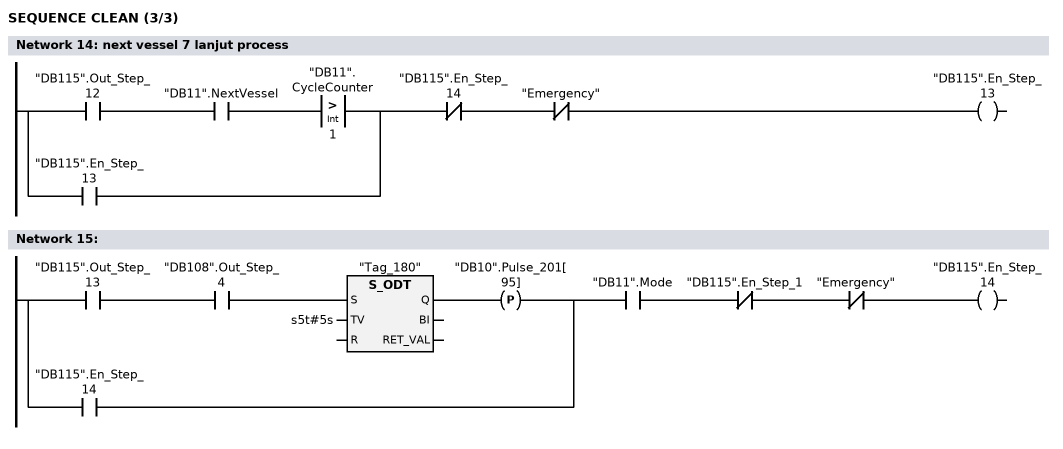
   RUNG wire#powerrail
      Contact( "DB115".Out_Step_12 )
      Contact( "DB11".NextVessel )
      { S7_Templates := "SrcType := Int" } GT_Contact(in1 := "DB11".CycleCounter, in2 := 1)
      wire#w1
      I_Contact( "DB115".En_Step_14 )
      I_Contact( "Emergency" )
      Coil( "DB115".En_Step_13 )
   END_RUNG
   RUNG wire#powerrail
      Contact( "DB115".En_Step_13 )
   END_RUNG wire#w1
   // the same network as SCL:
   "DB115".En_Step_13 := (("DB115".Out_Step_12 AND "DB11".NextVessel AND ("DB11".CycleCounter > 1)) OR "DB115".En_Step_13) AND NOT "DB115".En_Step_14 AND NOT "Emergency";
END_REGION

REGION Network 15
   RUNG wire#powerrail
      Contact( "DB115".Out_Step_13 )
      Contact( "DB108".Out_Step_4 )
      S_ODT(T_NO := "Tag_180", TV := s5t#5s, R :=, BI =>, RET_VAL =>)
      P_Trig( "DB10".Pulse_201[95] )
      wire#w1
      Contact( "DB11".Mode )
      I_Contact( "DB115".En_Step_1 )
      I_Contact( "Emergency" )
      Coil( "DB115".En_Step_14 )
   END_RUNG
   RUNG wire#powerrail
      Contact( "DB115".En_Step_14 )
   END_RUNG wire#w1
   // the same network as SCL:
   #_s5time1 := S_ODT(T_NO := "Tag_180",
                      S := "DB115".Out_Step_13 AND "DB108".Out_Step_4,
                      TV := s5t#5s,
                      Q => #_w1);
   #_w2 := #_w1 AND NOT "DB10".Pulse_201[95];   // rising edge
   "DB10".Pulse_201[95] := #_w1;
   "DB115".En_Step_14 := (#_w2 OR "DB115".En_Step_14) AND "DB11".Mode AND NOT "DB115".En_Step_1 AND NOT "Emergency";
END_REGION
END_FUNCTION

FUNCTION "SEQUENCE CYCLE" : Void   // FC36, LAD
{ S7_Optimized_Access := 'TRUE' }
VERSION : 0.1
   VAR_TEMP   // added for the SCL form of the ladder/FBD networks
      _w1 : Bool;
      _w2 : Bool;
      _w3 : Bool;
      _s5time1 : S5Time;
      _w4 : Bool;
      _w5 : Bool;
   END_VAR
BEGIN

REGION Network 1: Dari supply ke vessel 1
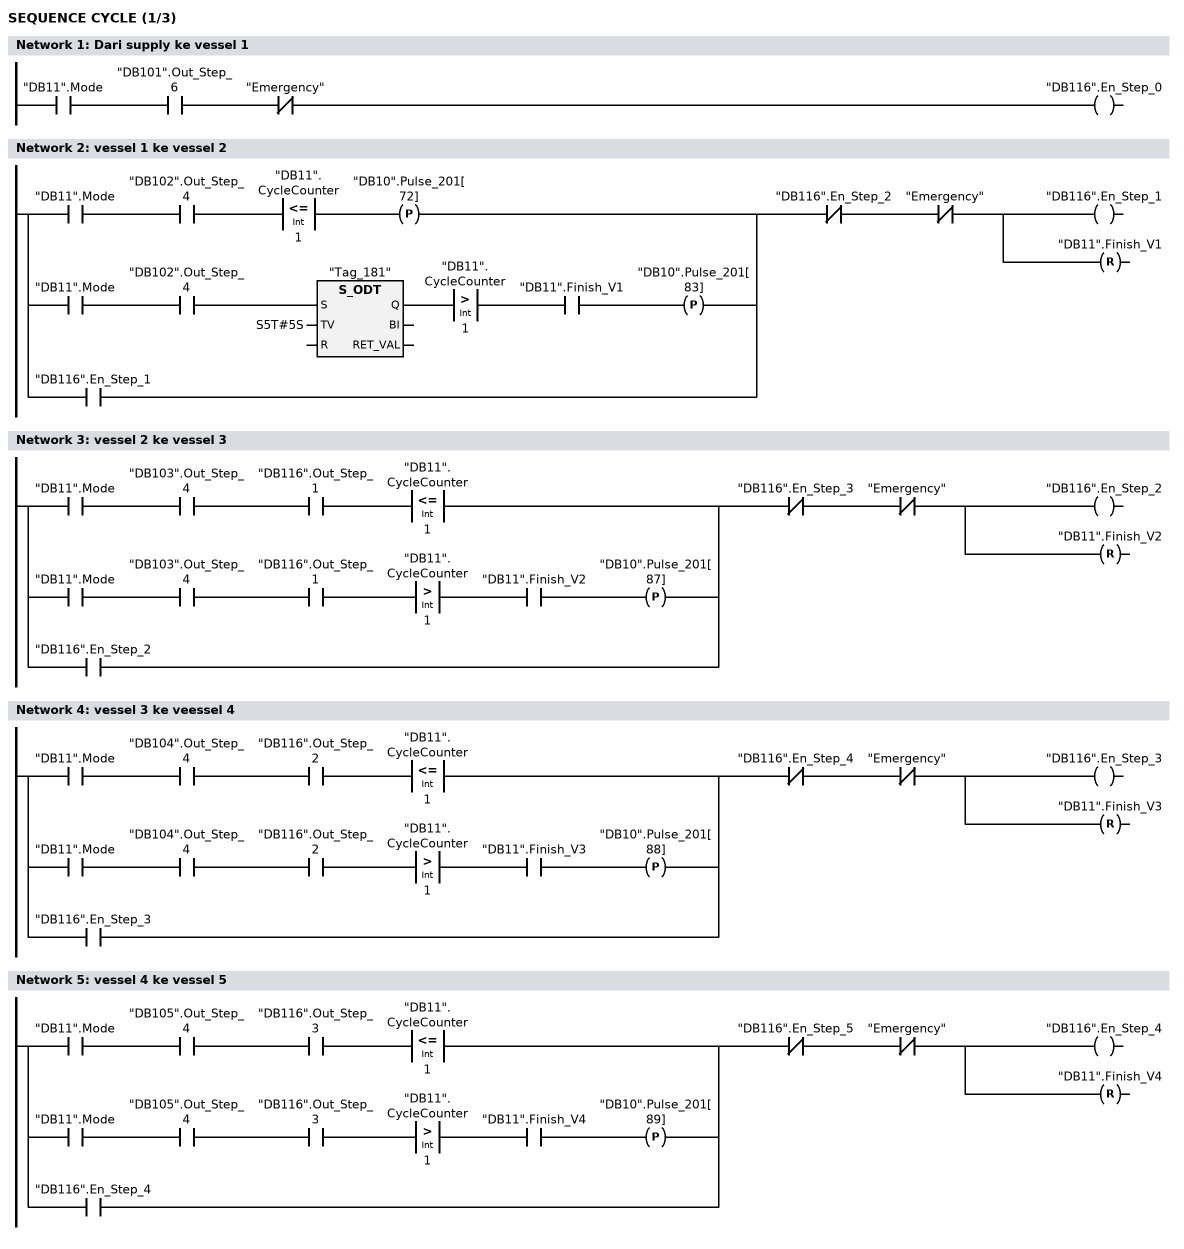
   RUNG wire#powerrail
      Contact( "DB11".Mode )
      Contact( "DB101".Out_Step_6 )
      I_Contact( "Emergency" )
      Coil( "DB116".En_Step_0 )
   END_RUNG
   // the same network as SCL:
   "DB116".En_Step_0 := "DB11".Mode AND "DB101".Out_Step_6 AND NOT "Emergency";
END_REGION

REGION Network 2: vessel 1 ke vessel 2
   RUNG wire#powerrail
      Contact( "DB11".Mode )
      Contact( "DB102".Out_Step_4 )
      { S7_Templates := "SrcType := Int" } LE_Contact(in1 := "DB11".CycleCounter, in2 := 1)
      P_Trig( "DB10".Pulse_201[72] )
      wire#w1
      I_Contact( "DB116".En_Step_2 )
      I_Contact( "Emergency" )
      wire#w2
      Coil( "DB116".En_Step_1 )
   END_RUNG
   RUNG wire#powerrail
      Contact( "DB11".Mode )
      Contact( "DB102".Out_Step_4 )
      S_ODT(T_NO := "Tag_181", TV := S5T#5S, R :=, BI =>, RET_VAL =>)
      { S7_Templates := "SrcType := Int" } GT_Contact(in1 := "DB11".CycleCounter, in2 := 1)
      Contact( "DB11".Finish_V1 )
      P_Trig( "DB10".Pulse_201[83] )
   END_RUNG wire#w1
   RUNG wire#powerrail
      Contact( "DB116".En_Step_1 )
   END_RUNG wire#w1
   RUNG wire#w2
      R_Coil( "DB11".Finish_V1 )
   END_RUNG
   // the same network as SCL:
   #_w1 := "DB11".Mode AND "DB102".Out_Step_4 AND ("DB11".CycleCounter <= 1);
   #_w2 := #_w1 AND NOT "DB10".Pulse_201[72];   // rising edge
   "DB10".Pulse_201[72] := #_w1;
   #_s5time1 := S_ODT(T_NO := "Tag_181", S := "DB11".Mode AND "DB102".Out_Step_4, TV := S5T#5S, Q => #_w3);
   #_w4 := #_w3 AND ("DB11".CycleCounter > 1) AND "DB11".Finish_V1;
   #_w5 := #_w4 AND NOT "DB10".Pulse_201[83];   // rising edge
   "DB10".Pulse_201[83] := #_w4;
   "DB116".En_Step_1 := (#_w2 OR #_w5 OR "DB116".En_Step_1) AND NOT "DB116".En_Step_2 AND NOT "Emergency";
   IF "DB116".En_Step_1 THEN "DB11".Finish_V1 := FALSE; END_IF;
END_REGION

REGION Network 3: vessel 2 ke vessel 3
   RUNG wire#powerrail
      Contact( "DB11".Mode )
      Contact( "DB103".Out_Step_4 )
      Contact( "DB116".Out_Step_1 )
      { S7_Templates := "SrcType := Int" } LE_Contact(in1 := "DB11".CycleCounter, in2 := 1)
      wire#w1
      I_Contact( "DB116".En_Step_3 )
      I_Contact( "Emergency" )
      wire#w2
      Coil( "DB116".En_Step_2 )
   END_RUNG
   RUNG wire#powerrail
      Contact( "DB11".Mode )
      Contact( "DB103".Out_Step_4 )
      Contact( "DB116".Out_Step_1 )
      { S7_Templates := "SrcType := Int" } GT_Contact(in1 := "DB11".CycleCounter, in2 := 1)
      Contact( "DB11".Finish_V2 )
      P_Trig( "DB10".Pulse_201[87] )
   END_RUNG wire#w1
   RUNG wire#powerrail
      Contact( "DB116".En_Step_2 )
   END_RUNG wire#w1
   RUNG wire#w2
      R_Coil( "DB11".Finish_V2 )
   END_RUNG
   // the same network as SCL:
   #_w1 := "DB11".Mode AND "DB103".Out_Step_4 AND "DB116".Out_Step_1 AND ("DB11".CycleCounter > 1) AND "DB11".Finish_V2;
   #_w2 := #_w1 AND NOT "DB10".Pulse_201[87];   // rising edge
   "DB10".Pulse_201[87] := #_w1;
   "DB116".En_Step_2 := (("DB11".Mode AND "DB103".Out_Step_4 AND "DB116".Out_Step_1 AND ("DB11".CycleCounter <= 1)) OR #_w2 OR "DB116".En_Step_2) AND NOT "DB116".En_Step_3 AND NOT "Emergency";
   IF "DB116".En_Step_2 THEN "DB11".Finish_V2 := FALSE; END_IF;
END_REGION

REGION Network 4: vessel 3 ke veessel 4
   RUNG wire#powerrail
      Contact( "DB11".Mode )
      Contact( "DB104".Out_Step_4 )
      Contact( "DB116".Out_Step_2 )
      { S7_Templates := "SrcType := Int" } LE_Contact(in1 := "DB11".CycleCounter, in2 := 1)
      wire#w1
      I_Contact( "DB116".En_Step_4 )
      I_Contact( "Emergency" )
      wire#w2
      Coil( "DB116".En_Step_3 )
   END_RUNG
   RUNG wire#powerrail
      Contact( "DB11".Mode )
      Contact( "DB104".Out_Step_4 )
      Contact( "DB116".Out_Step_2 )
      { S7_Templates := "SrcType := Int" } GT_Contact(in1 := "DB11".CycleCounter, in2 := 1)
      Contact( "DB11".Finish_V3 )
      P_Trig( "DB10".Pulse_201[88] )
   END_RUNG wire#w1
   RUNG wire#powerrail
      Contact( "DB116".En_Step_3 )
   END_RUNG wire#w1
   RUNG wire#w2
      R_Coil( "DB11".Finish_V3 )
   END_RUNG
   // the same network as SCL:
   #_w1 := "DB11".Mode AND "DB104".Out_Step_4 AND "DB116".Out_Step_2 AND ("DB11".CycleCounter > 1) AND "DB11".Finish_V3;
   #_w2 := #_w1 AND NOT "DB10".Pulse_201[88];   // rising edge
   "DB10".Pulse_201[88] := #_w1;
   "DB116".En_Step_3 := (("DB11".Mode AND "DB104".Out_Step_4 AND "DB116".Out_Step_2 AND ("DB11".CycleCounter <= 1)) OR #_w2 OR "DB116".En_Step_3) AND NOT "DB116".En_Step_4 AND NOT "Emergency";
   IF "DB116".En_Step_3 THEN "DB11".Finish_V3 := FALSE; END_IF;
END_REGION

REGION Network 5: vessel 4 ke vessel 5
   RUNG wire#powerrail
      Contact( "DB11".Mode )
      Contact( "DB105".Out_Step_4 )
      Contact( "DB116".Out_Step_3 )
      { S7_Templates := "SrcType := Int" } LE_Contact(in1 := "DB11".CycleCounter, in2 := 1)
      wire#w1
      I_Contact( "DB116".En_Step_5 )
      I_Contact( "Emergency" )
      wire#w2
      Coil( "DB116".En_Step_4 )
   END_RUNG
   RUNG wire#powerrail
      Contact( "DB11".Mode )
      Contact( "DB105".Out_Step_4 )
      Contact( "DB116".Out_Step_3 )
      { S7_Templates := "SrcType := Int" } GT_Contact(in1 := "DB11".CycleCounter, in2 := 1)
      Contact( "DB11".Finish_V4 )
      P_Trig( "DB10".Pulse_201[89] )
   END_RUNG wire#w1
   RUNG wire#powerrail
      Contact( "DB116".En_Step_4 )
   END_RUNG wire#w1
   RUNG wire#w2
      R_Coil( "DB11".Finish_V4 )
   END_RUNG
   // the same network as SCL:
   #_w1 := "DB11".Mode AND "DB105".Out_Step_4 AND "DB116".Out_Step_3 AND ("DB11".CycleCounter > 1) AND "DB11".Finish_V4;
   #_w2 := #_w1 AND NOT "DB10".Pulse_201[89];   // rising edge
   "DB10".Pulse_201[89] := #_w1;
   "DB116".En_Step_4 := (("DB11".Mode AND "DB105".Out_Step_4 AND "DB116".Out_Step_3 AND ("DB11".CycleCounter <= 1)) OR #_w2 OR "DB116".En_Step_4) AND NOT "DB116".En_Step_5 AND NOT "Emergency";
   IF "DB116".En_Step_4 THEN "DB11".Finish_V4 := FALSE; END_IF;
END_REGION

REGION Network 6: vessel 5 ke vessel 6
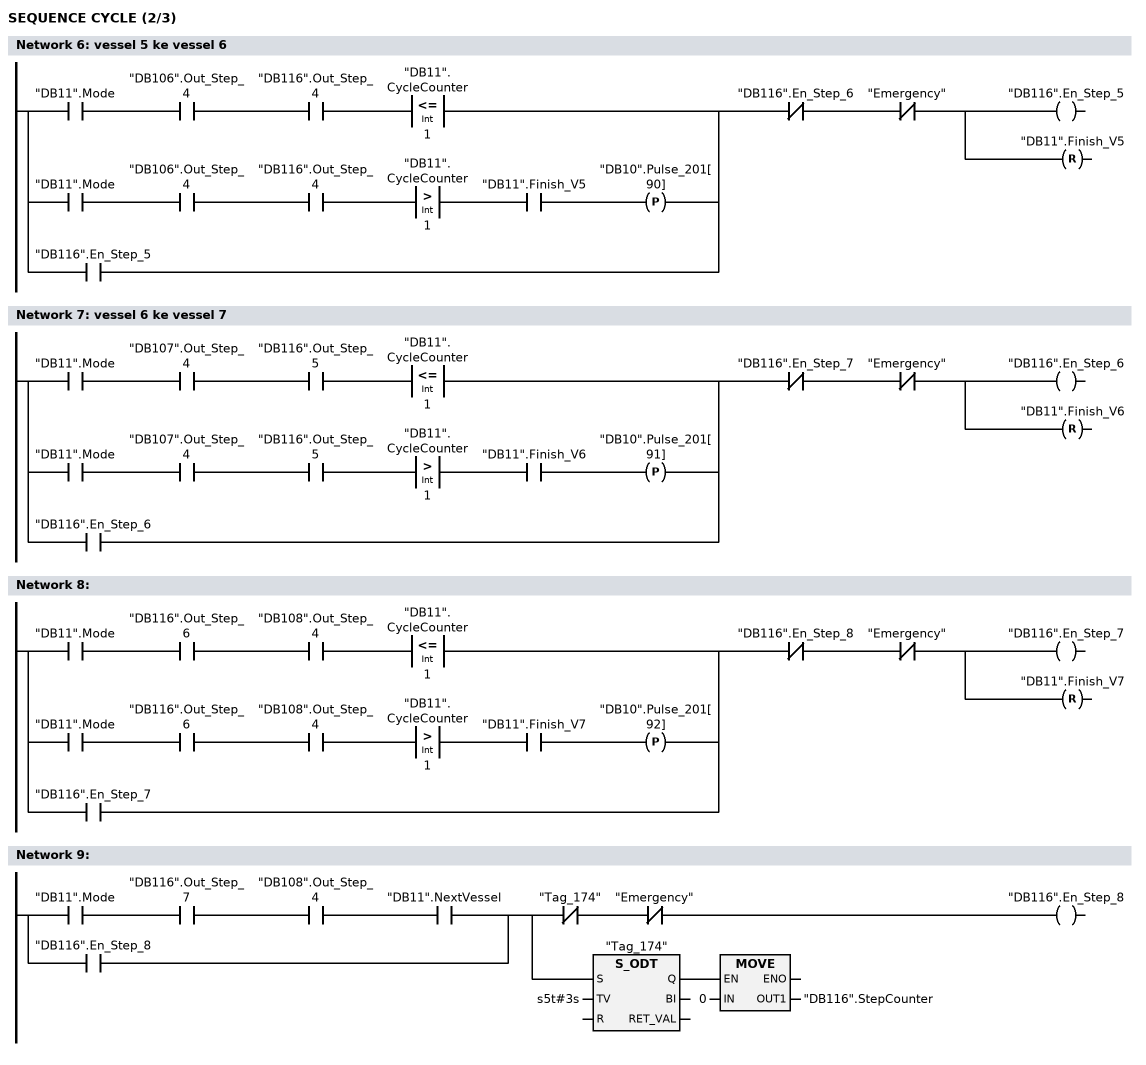
   RUNG wire#powerrail
      Contact( "DB11".Mode )
      Contact( "DB106".Out_Step_4 )
      Contact( "DB116".Out_Step_4 )
      { S7_Templates := "SrcType := Int" } LE_Contact(in1 := "DB11".CycleCounter, in2 := 1)
      wire#w1
      I_Contact( "DB116".En_Step_6 )
      I_Contact( "Emergency" )
      wire#w2
      Coil( "DB116".En_Step_5 )
   END_RUNG
   RUNG wire#powerrail
      Contact( "DB11".Mode )
      Contact( "DB106".Out_Step_4 )
      Contact( "DB116".Out_Step_4 )
      { S7_Templates := "SrcType := Int" } GT_Contact(in1 := "DB11".CycleCounter, in2 := 1)
      Contact( "DB11".Finish_V5 )
      P_Trig( "DB10".Pulse_201[90] )
   END_RUNG wire#w1
   RUNG wire#powerrail
      Contact( "DB116".En_Step_5 )
   END_RUNG wire#w1
   RUNG wire#w2
      R_Coil( "DB11".Finish_V5 )
   END_RUNG
   // the same network as SCL:
   #_w1 := "DB11".Mode AND "DB106".Out_Step_4 AND "DB116".Out_Step_4 AND ("DB11".CycleCounter > 1) AND "DB11".Finish_V5;
   #_w2 := #_w1 AND NOT "DB10".Pulse_201[90];   // rising edge
   "DB10".Pulse_201[90] := #_w1;
   "DB116".En_Step_5 := (("DB11".Mode AND "DB106".Out_Step_4 AND "DB116".Out_Step_4 AND ("DB11".CycleCounter <= 1)) OR #_w2 OR "DB116".En_Step_5) AND NOT "DB116".En_Step_6 AND NOT "Emergency";
   IF "DB116".En_Step_5 THEN "DB11".Finish_V5 := FALSE; END_IF;
END_REGION

REGION Network 7: vessel 6 ke vessel 7
   RUNG wire#powerrail
      Contact( "DB11".Mode )
      Contact( "DB107".Out_Step_4 )
      Contact( "DB116".Out_Step_5 )
      { S7_Templates := "SrcType := Int" } LE_Contact(in1 := "DB11".CycleCounter, in2 := 1)
      wire#w1
      I_Contact( "DB116".En_Step_7 )
      I_Contact( "Emergency" )
      wire#w2
      Coil( "DB116".En_Step_6 )
   END_RUNG
   RUNG wire#powerrail
      Contact( "DB11".Mode )
      Contact( "DB107".Out_Step_4 )
      Contact( "DB116".Out_Step_5 )
      { S7_Templates := "SrcType := Int" } GT_Contact(in1 := "DB11".CycleCounter, in2 := 1)
      Contact( "DB11".Finish_V6 )
      P_Trig( "DB10".Pulse_201[91] )
   END_RUNG wire#w1
   RUNG wire#powerrail
      Contact( "DB116".En_Step_6 )
   END_RUNG wire#w1
   RUNG wire#w2
      R_Coil( "DB11".Finish_V6 )
   END_RUNG
   // the same network as SCL:
   #_w1 := "DB11".Mode AND "DB107".Out_Step_4 AND "DB116".Out_Step_5 AND ("DB11".CycleCounter > 1) AND "DB11".Finish_V6;
   #_w2 := #_w1 AND NOT "DB10".Pulse_201[91];   // rising edge
   "DB10".Pulse_201[91] := #_w1;
   "DB116".En_Step_6 := (("DB11".Mode AND "DB107".Out_Step_4 AND "DB116".Out_Step_5 AND ("DB11".CycleCounter <= 1)) OR #_w2 OR "DB116".En_Step_6) AND NOT "DB116".En_Step_7 AND NOT "Emergency";
   IF "DB116".En_Step_6 THEN "DB11".Finish_V6 := FALSE; END_IF;
END_REGION

REGION Network 8
   RUNG wire#powerrail
      Contact( "DB11".Mode )
      Contact( "DB116".Out_Step_6 )
      Contact( "DB108".Out_Step_4 )
      { S7_Templates := "SrcType := Int" } LE_Contact(in1 := "DB11".CycleCounter, in2 := 1)
      wire#w1
      I_Contact( "DB116".En_Step_8 )
      I_Contact( "Emergency" )
      wire#w2
      Coil( "DB116".En_Step_7 )
   END_RUNG
   RUNG wire#powerrail
      Contact( "DB11".Mode )
      Contact( "DB116".Out_Step_6 )
      Contact( "DB108".Out_Step_4 )
      { S7_Templates := "SrcType := Int" } GT_Contact(in1 := "DB11".CycleCounter, in2 := 1)
      Contact( "DB11".Finish_V7 )
      P_Trig( "DB10".Pulse_201[92] )
   END_RUNG wire#w1
   RUNG wire#powerrail
      Contact( "DB116".En_Step_7 )
   END_RUNG wire#w1
   RUNG wire#w2
      R_Coil( "DB11".Finish_V7 )
   END_RUNG
   // the same network as SCL:
   #_w1 := "DB11".Mode AND "DB116".Out_Step_6 AND "DB108".Out_Step_4 AND ("DB11".CycleCounter > 1) AND "DB11".Finish_V7;
   #_w2 := #_w1 AND NOT "DB10".Pulse_201[92];   // rising edge
   "DB10".Pulse_201[92] := #_w1;
   "DB116".En_Step_7 := (("DB11".Mode AND "DB116".Out_Step_6 AND "DB108".Out_Step_4 AND ("DB11".CycleCounter <= 1)) OR #_w2 OR "DB116".En_Step_7) AND NOT "DB116".En_Step_8 AND NOT "Emergency";
   IF "DB116".En_Step_7 THEN "DB11".Finish_V7 := FALSE; END_IF;
END_REGION

REGION Network 9
   RUNG wire#powerrail
      Contact( "DB11".Mode )
      Contact( "DB116".Out_Step_7 )
      Contact( "DB108".Out_Step_4 )
      Contact( "DB11".NextVessel )
      wire#w1
      I_Contact( "Tag_174" )
      I_Contact( "Emergency" )
      Coil( "DB116".En_Step_8 )
   END_RUNG
   RUNG wire#powerrail
      Contact( "DB116".En_Step_8 )
   END_RUNG wire#w1
   RUNG wire#w1
      S_ODT(T_NO := "Tag_174", TV := s5t#3s, R :=, BI =>, RET_VAL =>)
      Move(in := 0, out1 => "DB116".StepCounter)
   END_RUNG
   // the same network as SCL:
   #_w1 := ("DB11".Mode AND "DB116".Out_Step_7 AND "DB108".Out_Step_4 AND "DB11".NextVessel) OR "DB116".En_Step_8;
   "DB116".En_Step_8 := #_w1 AND NOT "Tag_174" AND NOT "Emergency";
   #_s5time1 := S_ODT(T_NO := "Tag_174", S := #_w1, TV := s5t#3s, Q => #_w2);
   IF #_w2 THEN "DB116".StepCounter := 0; END_IF;
END_REGION

REGION Network 10
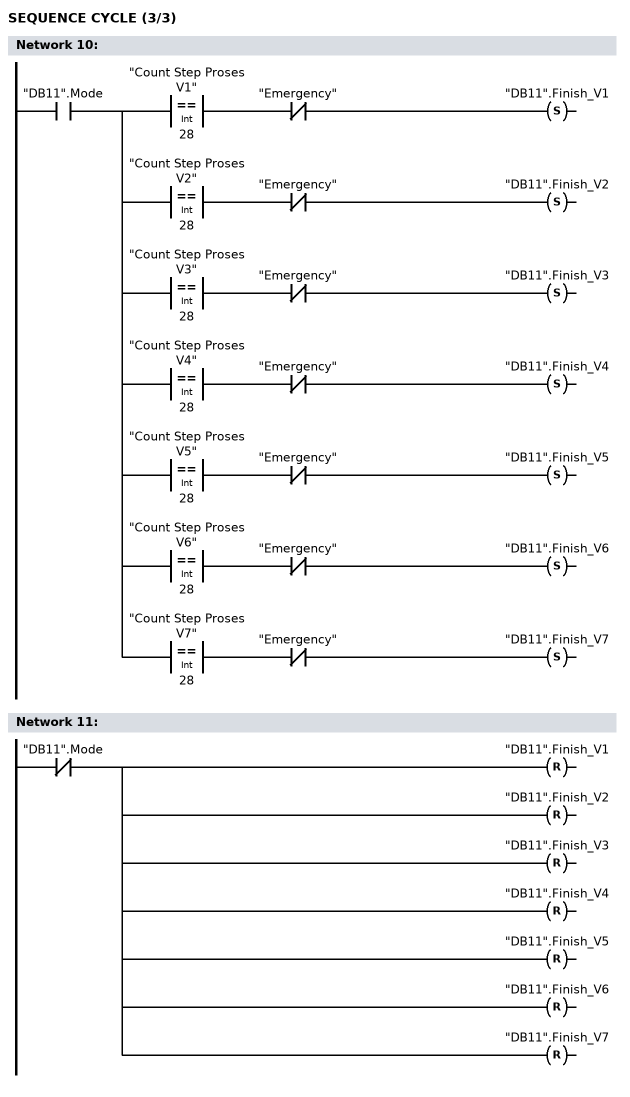
   RUNG wire#powerrail
      Contact( "DB11".Mode )
      wire#w1
      { S7_Templates := "SrcType := Int" } EQ_Contact(in1 := "Count Step Proses V1", in2 := 28)
      I_Contact( "Emergency" )
      S_Coil( "DB11".Finish_V1 )
   END_RUNG
   RUNG wire#w1
      { S7_Templates := "SrcType := Int" } EQ_Contact(in1 := "Count Step Proses V2", in2 := 28)
      I_Contact( "Emergency" )
      S_Coil( "DB11".Finish_V2 )
   END_RUNG
   RUNG wire#w1
      { S7_Templates := "SrcType := Int" } EQ_Contact(in1 := "Count Step Proses V3", in2 := 28)
      I_Contact( "Emergency" )
      S_Coil( "DB11".Finish_V3 )
   END_RUNG
   RUNG wire#w1
      { S7_Templates := "SrcType := Int" } EQ_Contact(in1 := "Count Step Proses V4", in2 := 28)
      I_Contact( "Emergency" )
      S_Coil( "DB11".Finish_V4 )
   END_RUNG
   RUNG wire#w1
      { S7_Templates := "SrcType := Int" } EQ_Contact(in1 := "Count Step Proses V5", in2 := 28)
      I_Contact( "Emergency" )
      S_Coil( "DB11".Finish_V5 )
   END_RUNG
   RUNG wire#w1
      { S7_Templates := "SrcType := Int" } EQ_Contact(in1 := "Count Step Proses V6", in2 := 28)
      I_Contact( "Emergency" )
      S_Coil( "DB11".Finish_V6 )
   END_RUNG
   RUNG wire#w1
      { S7_Templates := "SrcType := Int" } EQ_Contact(in1 := "Count Step Proses V7", in2 := 28)
      I_Contact( "Emergency" )
      S_Coil( "DB11".Finish_V7 )
   END_RUNG
   // the same network as SCL:
   IF "DB11".Mode AND ("Count Step Proses V1" = 28) AND NOT "Emergency" THEN
       "DB11".Finish_V1 := TRUE;
   END_IF;
   IF "DB11".Mode AND ("Count Step Proses V2" = 28) AND NOT "Emergency" THEN
       "DB11".Finish_V2 := TRUE;
   END_IF;
   IF "DB11".Mode AND ("Count Step Proses V3" = 28) AND NOT "Emergency" THEN
       "DB11".Finish_V3 := TRUE;
   END_IF;
   IF "DB11".Mode AND ("Count Step Proses V4" = 28) AND NOT "Emergency" THEN
       "DB11".Finish_V4 := TRUE;
   END_IF;
   IF "DB11".Mode AND ("Count Step Proses V5" = 28) AND NOT "Emergency" THEN
       "DB11".Finish_V5 := TRUE;
   END_IF;
   IF "DB11".Mode AND ("Count Step Proses V6" = 28) AND NOT "Emergency" THEN
       "DB11".Finish_V6 := TRUE;
   END_IF;
   IF "DB11".Mode AND ("Count Step Proses V7" = 28) AND NOT "Emergency" THEN
       "DB11".Finish_V7 := TRUE;
   END_IF;
END_REGION

REGION Network 11
   RUNG wire#powerrail
      I_Contact( "DB11".Mode )
      wire#w1
      R_Coil( "DB11".Finish_V1 )
   END_RUNG
   RUNG wire#w1
      R_Coil( "DB11".Finish_V2 )
   END_RUNG
   RUNG wire#w1
      R_Coil( "DB11".Finish_V3 )
   END_RUNG
   RUNG wire#w1
      R_Coil( "DB11".Finish_V4 )
   END_RUNG
   RUNG wire#w1
      R_Coil( "DB11".Finish_V5 )
   END_RUNG
   RUNG wire#w1
      R_Coil( "DB11".Finish_V6 )
   END_RUNG
   RUNG wire#w1
      R_Coil( "DB11".Finish_V7 )
   END_RUNG
   // the same network as SCL:
   IF NOT "DB11".Mode THEN
       "DB11".Finish_V1 := FALSE;
       "DB11".Finish_V2 := FALSE;
       "DB11".Finish_V3 := FALSE;
       "DB11".Finish_V4 := FALSE;
       "DB11".Finish_V5 := FALSE;
       "DB11".Finish_V6 := FALSE;
       "DB11".Finish_V7 := FALSE;
   END_IF;
END_REGION
END_FUNCTION

ORGANIZATION_BLOCK "Main"   // OB1, LAD, ProgramCycle
TITLE = "Main Program Sweep (Cycle)"
{ S7_Optimized_Access := 'TRUE' }
VERSION : 0.1
   VAR_INPUT
      Initial_Call : Bool;   // Initial call of this OB
      Remanence : Bool;   // =True, if remanent data are available
   END_VAR
   VAR_TEMP   // added for the SCL form of the ladder/FBD networks
      _w1 : Bool;
   END_VAR
BEGIN

REGION Network 1: PREPARATION VESSEL 1
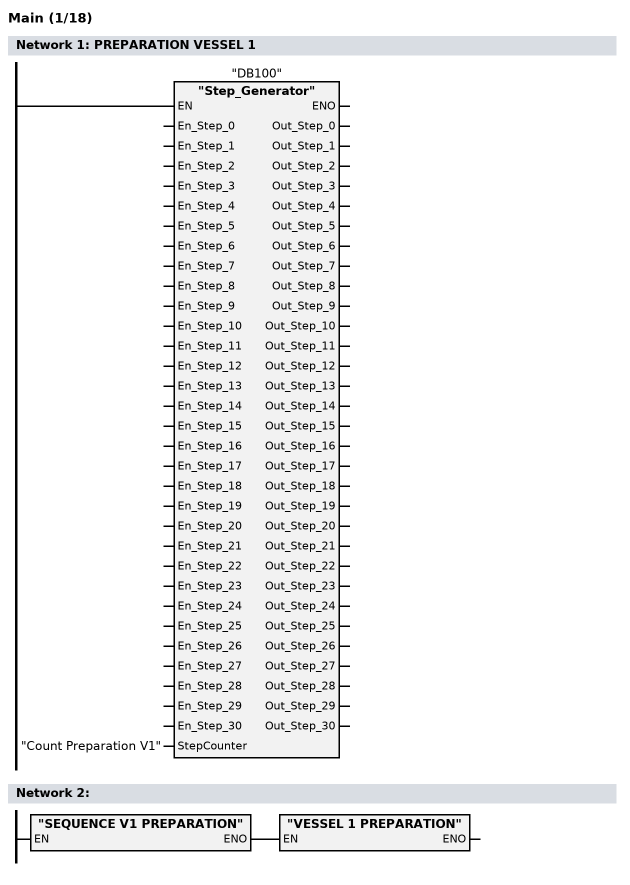
   RUNG wire#powerrail
      "DB100"(En_Step_0 :=, En_Step_1 :=, En_Step_2 :=, En_Step_3 :=, En_Step_4 :=, En_Step_5 :=, En_Step_6 :=, En_Step_7 :=, En_Step_8 :=, En_Step_9 :=, En_Step_10 :=, En_Step_11 :=, En_Step_12 :=, En_Step_13 :=, En_Step_14 :=, En_Step_15 :=, En_Step_16 :=, En_Step_17 :=, En_Step_18 :=, En_Step_19 :=, En_Step_20 :=, En_Step_21 :=, En_Step_22 :=, En_Step_23 :=, En_Step_24 :=, En_Step_25 :=, En_Step_26 :=, En_Step_27 :=, En_Step_28 :=, En_Step_29 :=, En_Step_30 :=, StepCounter := "Count Preparation V1", Out_Step_0 =>, Out_Step_1 =>, Out_Step_2 =>, Out_Step_3 =>, Out_Step_4 =>, Out_Step_5 =>, Out_Step_6 =>, Out_Step_7 =>, Out_Step_8 =>, Out_Step_9 =>, Out_Step_10 =>, Out_Step_11 =>, Out_Step_12 =>, Out_Step_13 =>, Out_Step_14 =>, Out_Step_15 =>, Out_Step_16 =>, Out_Step_17 =>, Out_Step_18 =>, Out_Step_19 =>, Out_Step_20 =>, Out_Step_21 =>, Out_Step_22 =>, Out_Step_23 =>, Out_Step_24 =>, Out_Step_25 =>, Out_Step_26 =>, Out_Step_27 =>, Out_Step_28 =>, Out_Step_29 =>, Out_Step_30 =>)
   END_RUNG
   // the same network as SCL:
   "DB100"(StepCounter := "Count Preparation V1");   // "Step_Generator"
END_REGION

REGION Network 2
   RUNG wire#powerrail
      "SEQUENCE V1 PREPARATION"()
      "VESSEL 1 PREPARATION"()
   END_RUNG
   // the same network as SCL:
   "SEQUENCE V1 PREPARATION"(ENO => #_w1);
   IF #_w1 THEN "VESSEL 1 PREPARATION"(); END_IF;
END_REGION

REGION Network 3: PREPARATION VESSEL 2
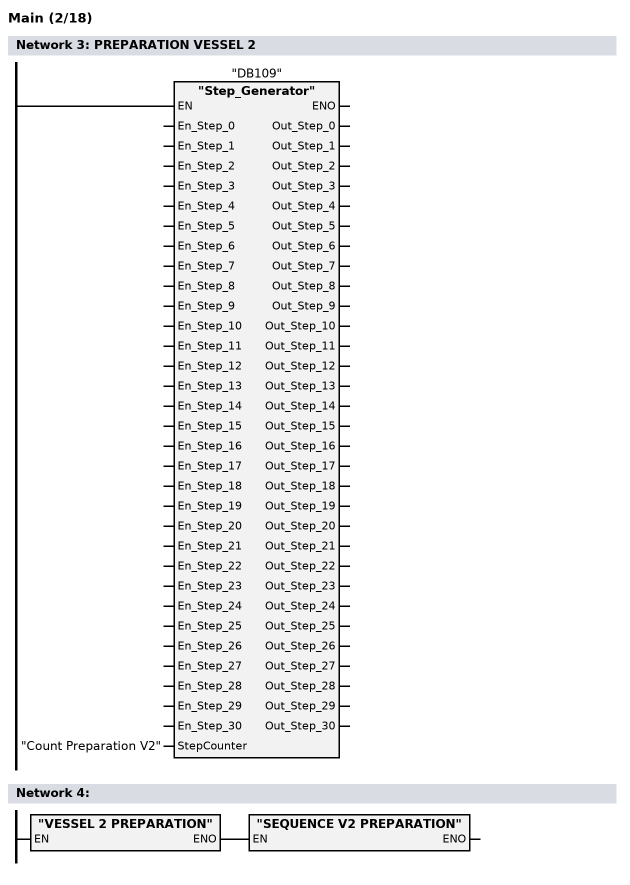
   RUNG wire#powerrail
      "DB109"(En_Step_0 :=, En_Step_1 :=, En_Step_2 :=, En_Step_3 :=, En_Step_4 :=, En_Step_5 :=, En_Step_6 :=, En_Step_7 :=, En_Step_8 :=, En_Step_9 :=, En_Step_10 :=, En_Step_11 :=, En_Step_12 :=, En_Step_13 :=, En_Step_14 :=, En_Step_15 :=, En_Step_16 :=, En_Step_17 :=, En_Step_18 :=, En_Step_19 :=, En_Step_20 :=, En_Step_21 :=, En_Step_22 :=, En_Step_23 :=, En_Step_24 :=, En_Step_25 :=, En_Step_26 :=, En_Step_27 :=, En_Step_28 :=, En_Step_29 :=, En_Step_30 :=, StepCounter := "Count Preparation V2", Out_Step_0 =>, Out_Step_1 =>, Out_Step_2 =>, Out_Step_3 =>, Out_Step_4 =>, Out_Step_5 =>, Out_Step_6 =>, Out_Step_7 =>, Out_Step_8 =>, Out_Step_9 =>, Out_Step_10 =>, Out_Step_11 =>, Out_Step_12 =>, Out_Step_13 =>, Out_Step_14 =>, Out_Step_15 =>, Out_Step_16 =>, Out_Step_17 =>, Out_Step_18 =>, Out_Step_19 =>, Out_Step_20 =>, Out_Step_21 =>, Out_Step_22 =>, Out_Step_23 =>, Out_Step_24 =>, Out_Step_25 =>, Out_Step_26 =>, Out_Step_27 =>, Out_Step_28 =>, Out_Step_29 =>, Out_Step_30 =>)
   END_RUNG
   // the same network as SCL:
   "DB109"(StepCounter := "Count Preparation V2");   // "Step_Generator"
END_REGION

REGION Network 4
   RUNG wire#powerrail
      "VESSEL 2 PREPARATION"()
      "SEQUENCE V2 PREPARATION"()
   END_RUNG
   // the same network as SCL:
   "VESSEL 2 PREPARATION"(ENO => #_w1);
   IF #_w1 THEN "SEQUENCE V2 PREPARATION"(); END_IF;
END_REGION

REGION Network 5: PREPARATION VESSEL 3
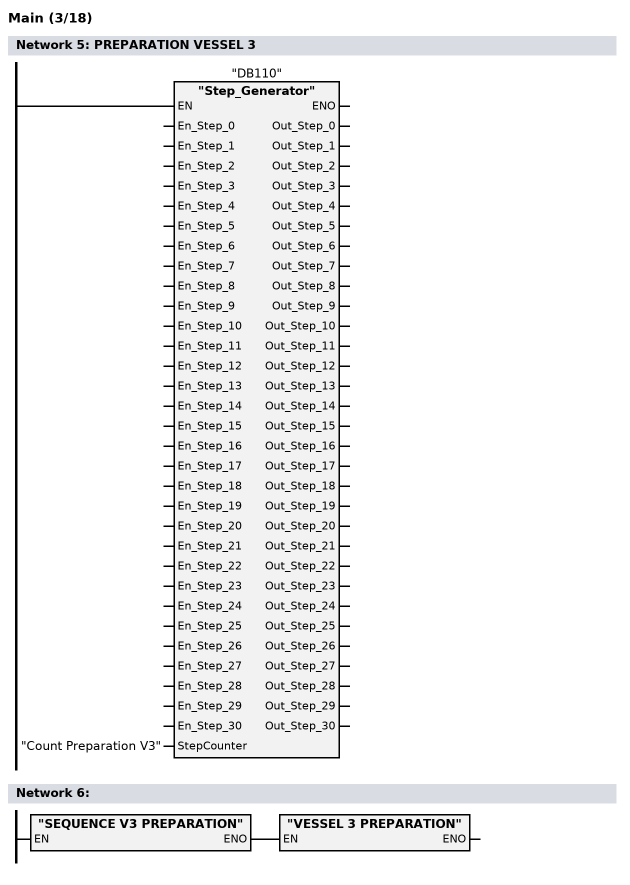
   RUNG wire#powerrail
      "DB110"(En_Step_0 :=, En_Step_1 :=, En_Step_2 :=, En_Step_3 :=, En_Step_4 :=, En_Step_5 :=, En_Step_6 :=, En_Step_7 :=, En_Step_8 :=, En_Step_9 :=, En_Step_10 :=, En_Step_11 :=, En_Step_12 :=, En_Step_13 :=, En_Step_14 :=, En_Step_15 :=, En_Step_16 :=, En_Step_17 :=, En_Step_18 :=, En_Step_19 :=, En_Step_20 :=, En_Step_21 :=, En_Step_22 :=, En_Step_23 :=, En_Step_24 :=, En_Step_25 :=, En_Step_26 :=, En_Step_27 :=, En_Step_28 :=, En_Step_29 :=, En_Step_30 :=, StepCounter := "Count Preparation V3", Out_Step_0 =>, Out_Step_1 =>, Out_Step_2 =>, Out_Step_3 =>, Out_Step_4 =>, Out_Step_5 =>, Out_Step_6 =>, Out_Step_7 =>, Out_Step_8 =>, Out_Step_9 =>, Out_Step_10 =>, Out_Step_11 =>, Out_Step_12 =>, Out_Step_13 =>, Out_Step_14 =>, Out_Step_15 =>, Out_Step_16 =>, Out_Step_17 =>, Out_Step_18 =>, Out_Step_19 =>, Out_Step_20 =>, Out_Step_21 =>, Out_Step_22 =>, Out_Step_23 =>, Out_Step_24 =>, Out_Step_25 =>, Out_Step_26 =>, Out_Step_27 =>, Out_Step_28 =>, Out_Step_29 =>, Out_Step_30 =>)
   END_RUNG
   // the same network as SCL:
   "DB110"(StepCounter := "Count Preparation V3");   // "Step_Generator"
END_REGION

REGION Network 6
   RUNG wire#powerrail
      "SEQUENCE V3 PREPARATION"()
      "VESSEL 3 PREPARATION"()
   END_RUNG
   // the same network as SCL:
   "SEQUENCE V3 PREPARATION"(ENO => #_w1);
   IF #_w1 THEN "VESSEL 3 PREPARATION"(); END_IF;
END_REGION

REGION Network 7: PREPARATION VESSEL 4
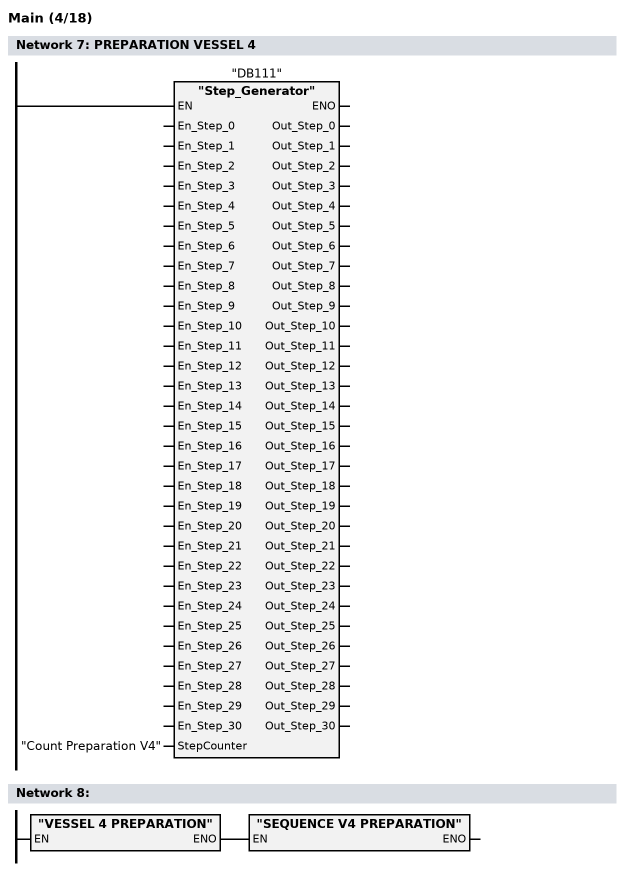
   RUNG wire#powerrail
      "DB111"(En_Step_0 :=, En_Step_1 :=, En_Step_2 :=, En_Step_3 :=, En_Step_4 :=, En_Step_5 :=, En_Step_6 :=, En_Step_7 :=, En_Step_8 :=, En_Step_9 :=, En_Step_10 :=, En_Step_11 :=, En_Step_12 :=, En_Step_13 :=, En_Step_14 :=, En_Step_15 :=, En_Step_16 :=, En_Step_17 :=, En_Step_18 :=, En_Step_19 :=, En_Step_20 :=, En_Step_21 :=, En_Step_22 :=, En_Step_23 :=, En_Step_24 :=, En_Step_25 :=, En_Step_26 :=, En_Step_27 :=, En_Step_28 :=, En_Step_29 :=, En_Step_30 :=, StepCounter := "Count Preparation V4", Out_Step_0 =>, Out_Step_1 =>, Out_Step_2 =>, Out_Step_3 =>, Out_Step_4 =>, Out_Step_5 =>, Out_Step_6 =>, Out_Step_7 =>, Out_Step_8 =>, Out_Step_9 =>, Out_Step_10 =>, Out_Step_11 =>, Out_Step_12 =>, Out_Step_13 =>, Out_Step_14 =>, Out_Step_15 =>, Out_Step_16 =>, Out_Step_17 =>, Out_Step_18 =>, Out_Step_19 =>, Out_Step_20 =>, Out_Step_21 =>, Out_Step_22 =>, Out_Step_23 =>, Out_Step_24 =>, Out_Step_25 =>, Out_Step_26 =>, Out_Step_27 =>, Out_Step_28 =>, Out_Step_29 =>, Out_Step_30 =>)
   END_RUNG
   // the same network as SCL:
   "DB111"(StepCounter := "Count Preparation V4");   // "Step_Generator"
END_REGION

REGION Network 8
   RUNG wire#powerrail
      "VESSEL 4 PREPARATION"()
      "SEQUENCE V4 PREPARATION"()
   END_RUNG
   // the same network as SCL:
   "VESSEL 4 PREPARATION"(ENO => #_w1);
   IF #_w1 THEN "SEQUENCE V4 PREPARATION"(); END_IF;
END_REGION

REGION Network 9: VESSEL 5 PREPARATION
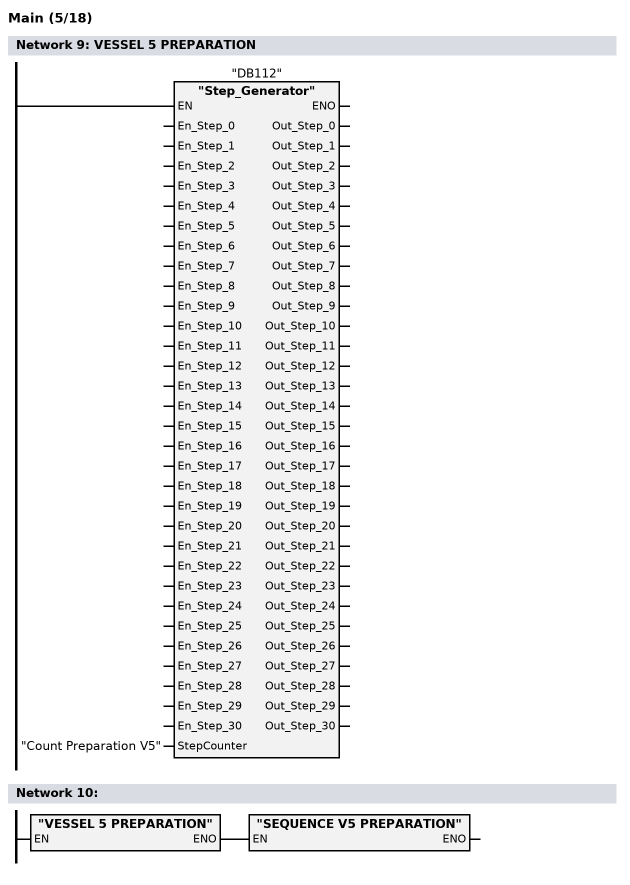
   RUNG wire#powerrail
      "DB112"(En_Step_0 :=, En_Step_1 :=, En_Step_2 :=, En_Step_3 :=, En_Step_4 :=, En_Step_5 :=, En_Step_6 :=, En_Step_7 :=, En_Step_8 :=, En_Step_9 :=, En_Step_10 :=, En_Step_11 :=, En_Step_12 :=, En_Step_13 :=, En_Step_14 :=, En_Step_15 :=, En_Step_16 :=, En_Step_17 :=, En_Step_18 :=, En_Step_19 :=, En_Step_20 :=, En_Step_21 :=, En_Step_22 :=, En_Step_23 :=, En_Step_24 :=, En_Step_25 :=, En_Step_26 :=, En_Step_27 :=, En_Step_28 :=, En_Step_29 :=, En_Step_30 :=, StepCounter := "Count Preparation V5", Out_Step_0 =>, Out_Step_1 =>, Out_Step_2 =>, Out_Step_3 =>, Out_Step_4 =>, Out_Step_5 =>, Out_Step_6 =>, Out_Step_7 =>, Out_Step_8 =>, Out_Step_9 =>, Out_Step_10 =>, Out_Step_11 =>, Out_Step_12 =>, Out_Step_13 =>, Out_Step_14 =>, Out_Step_15 =>, Out_Step_16 =>, Out_Step_17 =>, Out_Step_18 =>, Out_Step_19 =>, Out_Step_20 =>, Out_Step_21 =>, Out_Step_22 =>, Out_Step_23 =>, Out_Step_24 =>, Out_Step_25 =>, Out_Step_26 =>, Out_Step_27 =>, Out_Step_28 =>, Out_Step_29 =>, Out_Step_30 =>)
   END_RUNG
   // the same network as SCL:
   "DB112"(StepCounter := "Count Preparation V5");   // "Step_Generator"
END_REGION

REGION Network 10
   RUNG wire#powerrail
      "VESSEL 5 PREPARATION"()
      "SEQUENCE V5 PREPARATION"()
   END_RUNG
   // the same network as SCL:
   "VESSEL 5 PREPARATION"(ENO => #_w1);
   IF #_w1 THEN "SEQUENCE V5 PREPARATION"(); END_IF;
END_REGION

REGION Network 11: VESSEL 6 PREPARATION
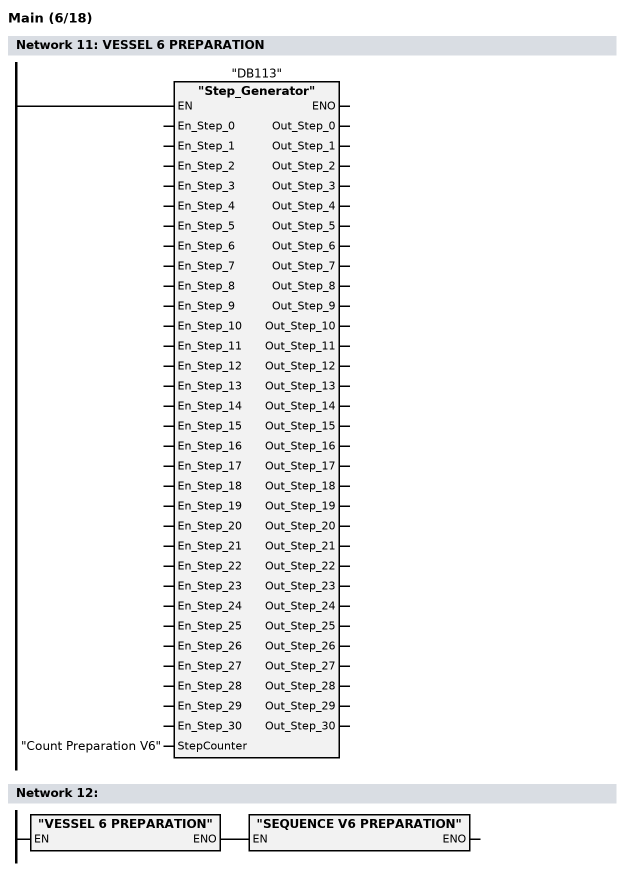
   RUNG wire#powerrail
      "DB113"(En_Step_0 :=, En_Step_1 :=, En_Step_2 :=, En_Step_3 :=, En_Step_4 :=, En_Step_5 :=, En_Step_6 :=, En_Step_7 :=, En_Step_8 :=, En_Step_9 :=, En_Step_10 :=, En_Step_11 :=, En_Step_12 :=, En_Step_13 :=, En_Step_14 :=, En_Step_15 :=, En_Step_16 :=, En_Step_17 :=, En_Step_18 :=, En_Step_19 :=, En_Step_20 :=, En_Step_21 :=, En_Step_22 :=, En_Step_23 :=, En_Step_24 :=, En_Step_25 :=, En_Step_26 :=, En_Step_27 :=, En_Step_28 :=, En_Step_29 :=, En_Step_30 :=, StepCounter := "Count Preparation V6", Out_Step_0 =>, Out_Step_1 =>, Out_Step_2 =>, Out_Step_3 =>, Out_Step_4 =>, Out_Step_5 =>, Out_Step_6 =>, Out_Step_7 =>, Out_Step_8 =>, Out_Step_9 =>, Out_Step_10 =>, Out_Step_11 =>, Out_Step_12 =>, Out_Step_13 =>, Out_Step_14 =>, Out_Step_15 =>, Out_Step_16 =>, Out_Step_17 =>, Out_Step_18 =>, Out_Step_19 =>, Out_Step_20 =>, Out_Step_21 =>, Out_Step_22 =>, Out_Step_23 =>, Out_Step_24 =>, Out_Step_25 =>, Out_Step_26 =>, Out_Step_27 =>, Out_Step_28 =>, Out_Step_29 =>, Out_Step_30 =>)
   END_RUNG
   // the same network as SCL:
   "DB113"(StepCounter := "Count Preparation V6");   // "Step_Generator"
END_REGION

REGION Network 12
   RUNG wire#powerrail
      "VESSEL 6 PREPARATION"()
      "SEQUENCE V6 PREPARATION"()
   END_RUNG
   // the same network as SCL:
   "VESSEL 6 PREPARATION"(ENO => #_w1);
   IF #_w1 THEN "SEQUENCE V6 PREPARATION"(); END_IF;
END_REGION

REGION Network 13: VESSEL 7 PREPARATION
